   
   COP(M215_M1_DR_OUT_MAJ,M215_M1_DR_IN_MAJ,1);
   M215_M1_DR_IN_MAR.EN := M215_M1_DR_OUT_MAR.EN;
   M215_M1_DR_IN_MAR.PC := M215_M1_DR_OUT_MAR.PC;
   COP(M215_M1_DR_OUT_MAM,M215_M1_DR_IN_MAM,1);
   COP(M215_M1_DR_OUT_MAS,M215_M1_DR_IN_MAS,1);
   COP(M215_M1_DR_OUT_MRP,M215_M1_DR_IN_MRP,1);
   COP(M215_M1_DR_OUT_MCD,M215_M1_DR_IN_MCD,1);
   
   COP(M216_M1_DR_OUT_MAJ,M216_M1_DR_IN_MAJ,1);
   M216_M1_DR_IN_MAR.EN := M216_M1_DR_OUT_MAR.EN;
   M216_M1_DR_IN_MAR.PC := M216_M1_DR_OUT_MAR.PC;
   COP(M216_M1_DR_OUT_MAM,M216_M1_DR_IN_MAM,1);
   COP(M216_M1_DR_OUT_MAS,M216_M1_DR_IN_MAS,1);
   COP(M216_M1_DR_OUT_MRP,M216_M1_DR_IN_MRP,1);
   COP(M216_M1_DR_OUT_MCD,M216_M1_DR_IN_MCD,1);
   
   COP(M217_M1_DR_OUT_MAJ,M217_M1_DR_IN_MAJ,1);
   M217_M1_DR_IN_MAR.EN := M217_M1_DR_OUT_MAR.EN;
   M217_M1_DR_IN_MAR.PC := M217_M1_DR_OUT_MAR.PC;
   COP(M217_M1_DR_OUT_MAM,M217_M1_DR_IN_MAM,1);
   COP(M217_M1_DR_OUT_MAS,M217_M1_DR_IN_MAS,1);
   COP(M217_M1_DR_OUT_MRP,M217_M1_DR_IN_MRP,1);
   COP(M217_M1_DR_OUT_MCD,M217_M1_DR_IN_MCD,1);
   
   COP(M218_M1_DR_OUT_MAJ,M218_M1_DR_IN_MAJ,1);
   M218_M1_DR_IN_MAR.EN := M218_M1_DR_OUT_MAR.EN;
   M218_M1_DR_IN_MAR.PC := M218_M1_DR_OUT_MAR.PC;
   COP(M218_M1_DR_OUT_MAM,M218_M1_DR_IN_MAM,1);
   COP(M218_M1_DR_OUT_MAS,M218_M1_DR_IN_MAS,1);
   COP(M218_M1_DR_OUT_MRP,M218_M1_DR_IN_MRP,1);
   COP(M218_M1_DR_OUT_MCD,M218_M1_DR_IN_MCD,1);
   
   COP(M219_M1_DR_OUT_MAJ,M219_M1_DR_IN_MAJ,1);
   M219_M1_DR_IN_MAR.EN := M219_M1_DR_OUT_MAR.EN;
   M219_M1_DR_IN_MAR.PC := M219_M1_DR_OUT_MAR.PC;
   COP(M219_M1_DR_OUT_MAM,M219_M1_DR_IN_MAM,1);
   COP(M219_M1_DR_OUT_MAS,M219_M1_DR_IN_MAS,1);
   COP(M219_M1_DR_OUT_MRP,M219_M1_DR_IN_MRP,1);
   COP(M219_M1_DR_OUT_MCD,M219_M1_DR_IN_MCD,1);
   
   COP(M220_M1_DR_OUT_MAJ,M220_M1_DR_IN_MAJ,1);
   M220_M1_DR_IN_MAR.EN := M220_M1_DR_OUT_MAR.EN;
   M220_M1_DR_IN_MAR.PC := M220_M1_DR_OUT_MAR.PC;
   COP(M220_M1_DR_OUT_MAM,M220_M1_DR_IN_MAM,1);
   COP(M220_M1_DR_OUT_MAS,M220_M1_DR_IN_MAS,1);
   COP(M220_M1_DR_OUT_MRP,M220_M1_DR_IN_MRP,1);
   COP(M220_M1_DR_OUT_MCD,M220_M1_DR_IN_MCD,1);
   
   COP(M225_M1_DR_OUT_MAJ,M225_M1_DR_IN_MAJ,1);
   M225_M1_DR_IN_MAR.EN := M225_M1_DR_OUT_MAR.EN;
   M225_M1_DR_IN_MAR.PC := M225_M1_DR_OUT_MAR.PC;
   COP(M225_M1_DR_OUT_MAM,M225_M1_DR_IN_MAM,1);
   COP(M225_M1_DR_OUT_MAS,M225_M1_DR_IN_MAS,1);
   COP(M225_M1_DR_OUT_MRP,M225_M1_DR_IN_MRP,1);
   COP(M225_M1_DR_OUT_MCD,M225_M1_DR_IN_MCD,1);
   
END_ROUTINE

ROUTINE _101_LADDER   (* ladder *)
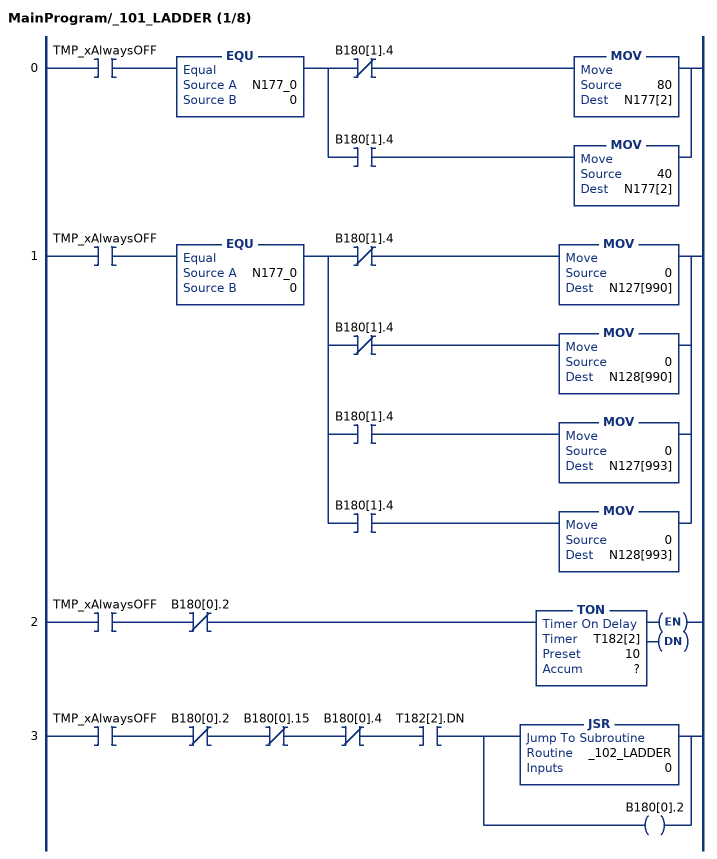
   0: XIC(TMP_xAlwaysOFF)EQU(N177_0,0)[XIO(B180[1].4) MOV(80,N177[2]) ,XIC(B180[1].4) MOV(40,N177[2]) ];
   1: XIC(TMP_xAlwaysOFF)EQU(N177_0,0)[XIO(B180[1].4) MOV(0,N127[990]) ,XIO(B180[1].4) MOV(0,N128[990]) ,XIC(B180[1].4) MOV(0,N127[993]) ,XIC(B180[1].4) MOV(0,N128[993]) ];
   2: XIC(TMP_xAlwaysOFF)XIO(B180[0].2)TON(T182[2],?,?);
   3: XIC(TMP_xAlwaysOFF)XIO(B180[0].2)XIO(B180[0].15)XIO(B180[0].4)XIC(T182[2].DN)[JSR(_102_LADDER,0) ,OTE(B180[0].2) ];
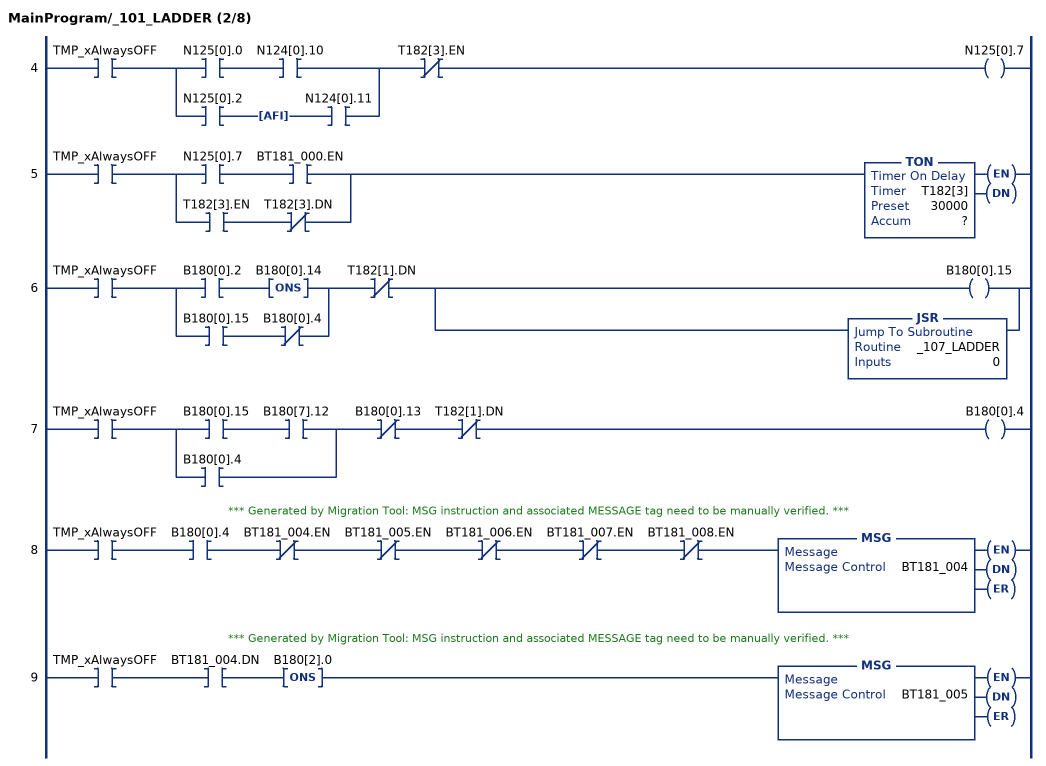
   4: XIC(TMP_xAlwaysOFF)[XIC(N125[0].0) XIC(N124[0].10) ,XIC(N125[0].2) AFI() XIC(N124[0].11) ]XIO(T182[3].EN)OTE(N125[0].7);
   5: XIC(TMP_xAlwaysOFF)[XIC(N125[0].7) XIC(BT181_000.EN) ,XIC(T182[3].EN) XIO(T182[3].DN) ]TON(T182[3],?,?);
   6: XIC(TMP_xAlwaysOFF)[XIC(B180[0].2) ONS(B180[0].14) ,XIC(B180[0].15) XIO(B180[0].4) ]XIO(T182[1].DN)[OTE(B180[0].15) ,JSR(_107_LADDER,0) ];
   7: XIC(TMP_xAlwaysOFF)[XIC(B180[0].15) XIC(B180[7].12) ,XIC(B180[0].4) ]XIO(B180[0].13)XIO(T182[1].DN)OTE(B180[0].4);
   // *** Generated by Migration Tool: MSG instruction and associated MESSAGE tag need to be manually verified. ***
   8: XIC(TMP_xAlwaysOFF)XIC(B180[0].4)XIO(BT181_004.EN)XIO(BT181_005.EN)XIO(BT181_006.EN)XIO(BT181_007.EN)XIO(BT181_008.EN)MSG(BT181_004);
   // *** Generated by Migration Tool: MSG instruction and associated MESSAGE tag need to be manually verified. ***
   9: XIC(TMP_xAlwaysOFF)XIC(BT181_004.DN)ONS(B180[2].0)MSG(BT181_005);
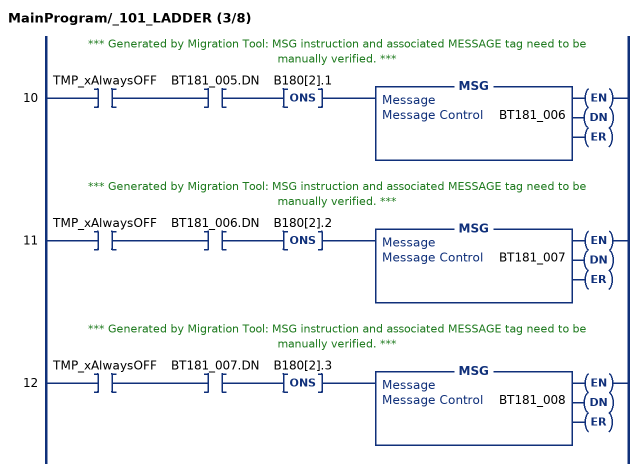
   // *** Generated by Migration Tool: MSG instruction and associated MESSAGE tag need to be manually verified. ***
   10: XIC(TMP_xAlwaysOFF)XIC(BT181_005.DN)ONS(B180[2].1)MSG(BT181_006);
   // *** Generated by Migration Tool: MSG instruction and associated MESSAGE tag need to be manually verified. ***
   11: XIC(TMP_xAlwaysOFF)XIC(BT181_006.DN)ONS(B180[2].2)MSG(BT181_007);
   // *** Generated by Migration Tool: MSG instruction and associated MESSAGE tag need to be manually verified. ***
   12: XIC(TMP_xAlwaysOFF)XIC(BT181_007.DN)ONS(B180[2].3)MSG(BT181_008);
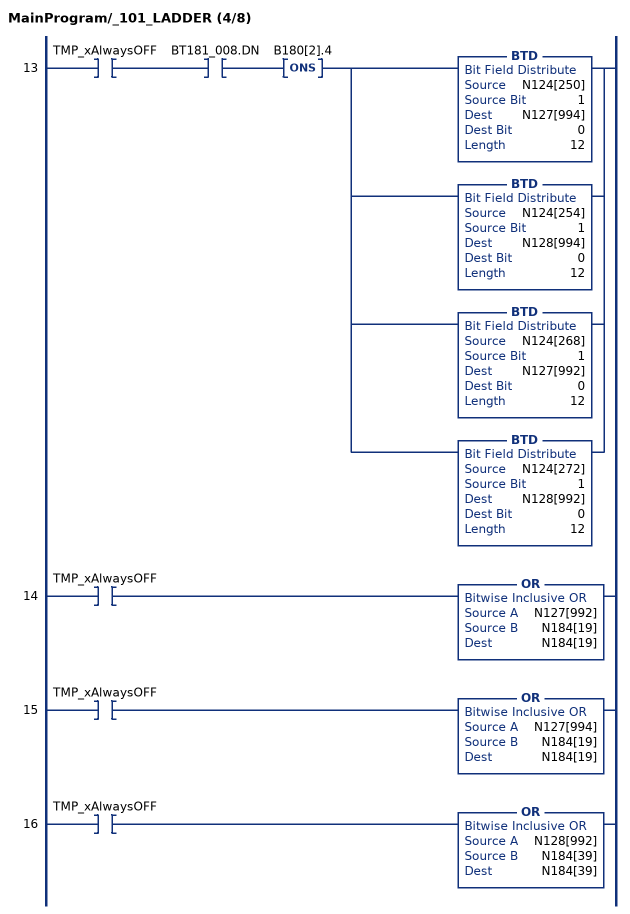
   13: XIC(TMP_xAlwaysOFF)XIC(BT181_008.DN)ONS(B180[2].4)[BTD(N124[250],1,N127[994],0,12) ,BTD(N124[254],1,N128[994],0,12) ,BTD(N124[268],1,N127[992],0,12) ,BTD(N124[272],1,N128[992],0,12) ];
   14: XIC(TMP_xAlwaysOFF)OR(N127[992],N184[19],N184[19]);
   15: XIC(TMP_xAlwaysOFF)OR(N127[994],N184[19],N184[19]);
   16: XIC(TMP_xAlwaysOFF)OR(N128[992],N184[39],N184[39]);
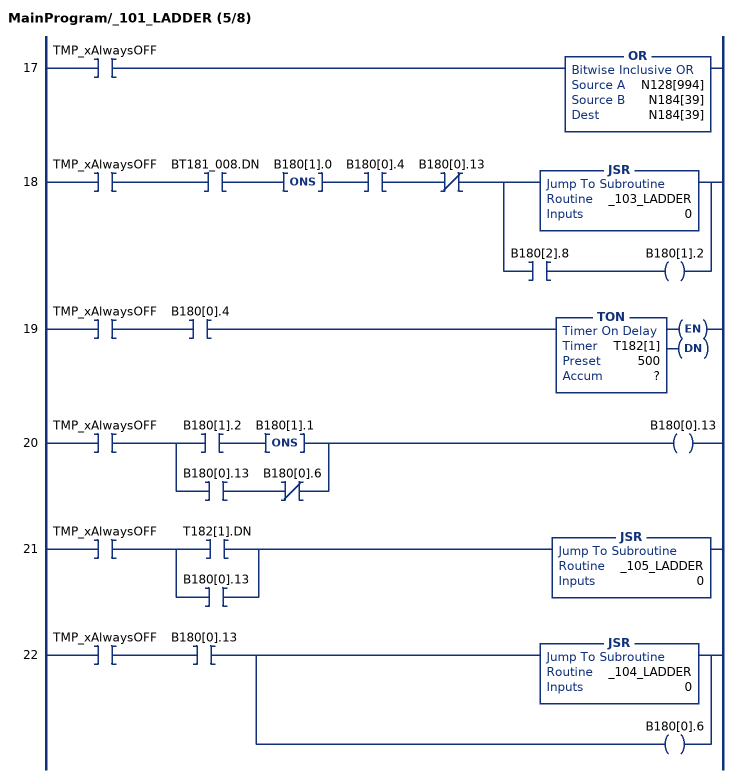
   17: XIC(TMP_xAlwaysOFF)OR(N128[994],N184[39],N184[39]);
   18: XIC(TMP_xAlwaysOFF)XIC(BT181_008.DN)ONS(B180[1].0)XIC(B180[0].4)XIO(B180[0].13)[JSR(_103_LADDER,0) ,XIC(B180[2].8) OTE(B180[1].2) ];
   19: XIC(TMP_xAlwaysOFF)XIC(B180[0].4)TON(T182[1],?,?);
   20: XIC(TMP_xAlwaysOFF)[XIC(B180[1].2) ONS(B180[1].1) ,XIC(B180[0].13) XIO(B180[0].6) ]OTE(B180[0].13);
   21: XIC(TMP_xAlwaysOFF)[XIC(T182[1].DN) ,XIC(B180[0].13) ]JSR(_105_LADDER,0);
   22: XIC(TMP_xAlwaysOFF)XIC(B180[0].13)[JSR(_104_LADDER,0) ,OTE(B180[0].6) ];
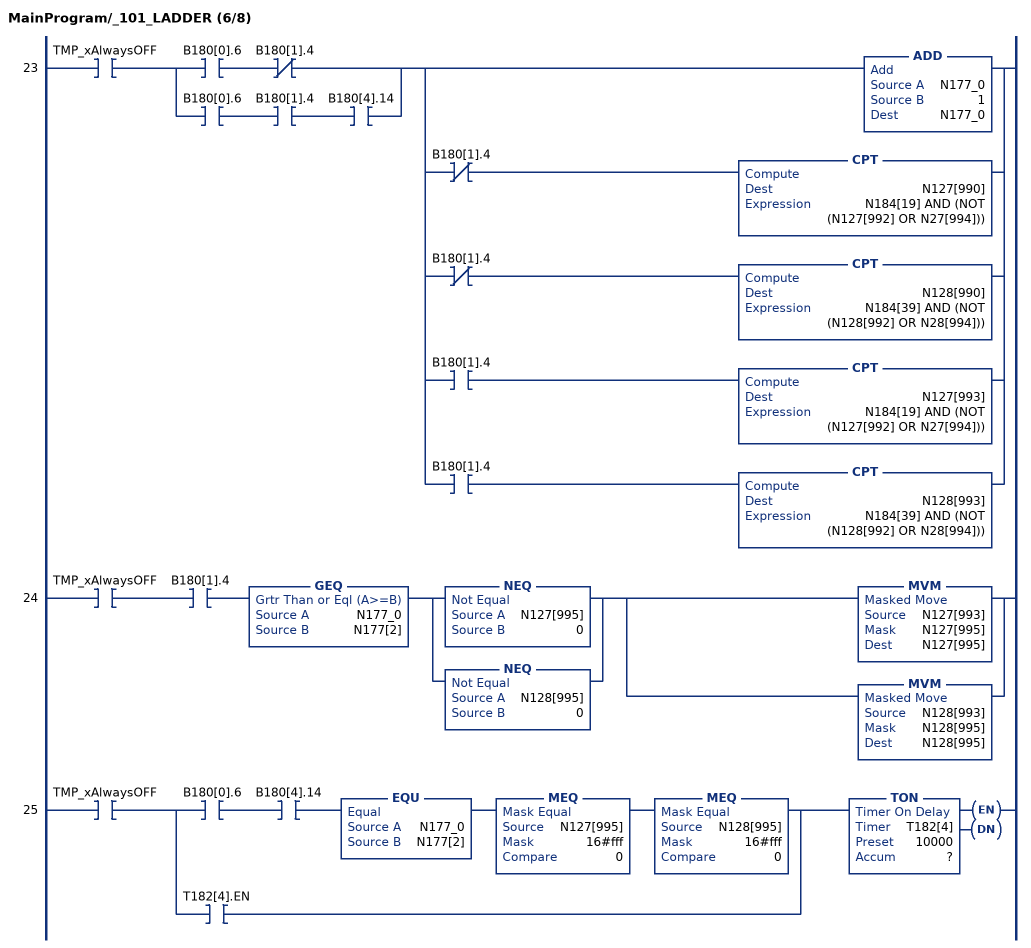
   23: XIC(TMP_xAlwaysOFF)[XIC(B180[0].6) XIO(B180[1].4) ,XIC(B180[0].6) XIC(B180[1].4) XIC(B180[4].14) ][ADD(N177_0,1,N177_0) ,XIO(B180[1].4) CPT(N127[990],N184[19] AND (NOT (N127[992] OR N27[994]))) ,XIO(B180[1].4) CPT(N128[990],N184[39] AND (NOT (N128[992] OR N28[994]))) ,XIC(B180[1].4) CPT(N127[993],N184[19] AND (NOT (N127[992] OR N27[994]))) ,XIC(B180[1].4) CPT(N128[993],N184[39] AND (NOT (N128[992] OR N28[994]))) ];
   24: XIC(TMP_xAlwaysOFF)XIC(B180[1].4)GEQ(N177_0,N177[2])[NEQ(N127[995],0) ,NEQ(N128[995],0) ][MVM(N127[993],N127[995],N127[995]) ,MVM(N128[993],N128[995],N128[995]) ];
   25: XIC(TMP_xAlwaysOFF)[XIC(B180[0].6) XIC(B180[4].14) EQU(N177_0,N177[2]) MEQ(N127[995],16#fff,0) MEQ(N128[995],16#fff,0) ,XIC(T182[4].EN) ]TON(T182[4],?,?);
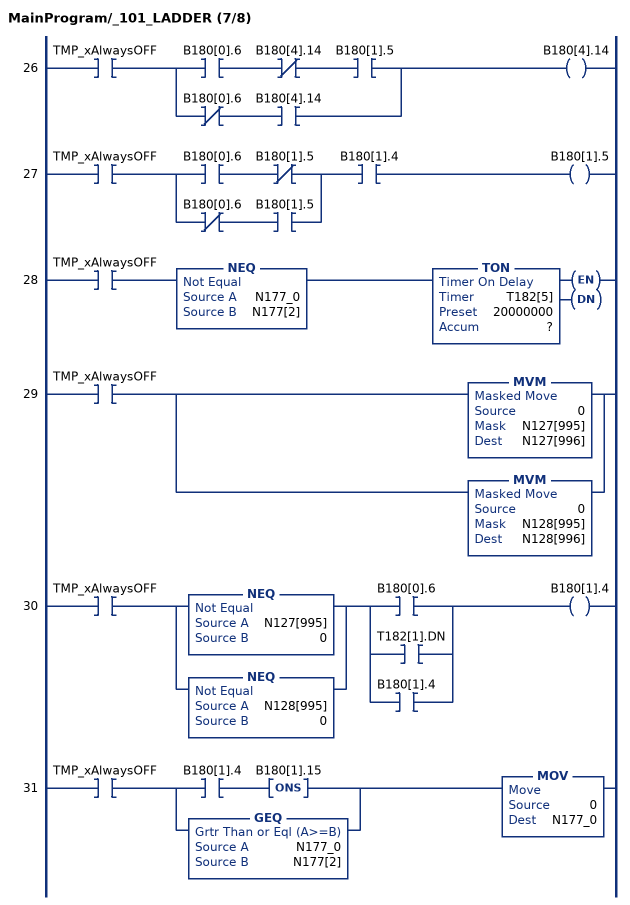
   26: XIC(TMP_xAlwaysOFF)[XIC(B180[0].6) XIO(B180[4].14) XIC(B180[1].5) ,XIO(B180[0].6) XIC(B180[4].14) ]OTE(B180[4].14);
   27: XIC(TMP_xAlwaysOFF)[XIC(B180[0].6) XIO(B180[1].5) ,XIO(B180[0].6) XIC(B180[1].5) ]XIC(B180[1].4)OTE(B180[1].5);
   28: XIC(TMP_xAlwaysOFF)NEQ(N177_0,N177[2])TON(T182[5],?,?);
   29: XIC(TMP_xAlwaysOFF)[MVM(0,N127[995],N127[996]) ,MVM(0,N128[995],N128[996]) ];
   30: XIC(TMP_xAlwaysOFF)[NEQ(N127[995],0) ,NEQ(N128[995],0) ][XIC(B180[0].6) ,XIC(T182[1].DN) ,XIC(B180[1].4) ]OTE(B180[1].4);
   31: XIC(TMP_xAlwaysOFF)[XIC(B180[1].4) ONS(B180[1].15) ,GEQ(N177_0,N177[2]) ]MOV(0,N177_0);
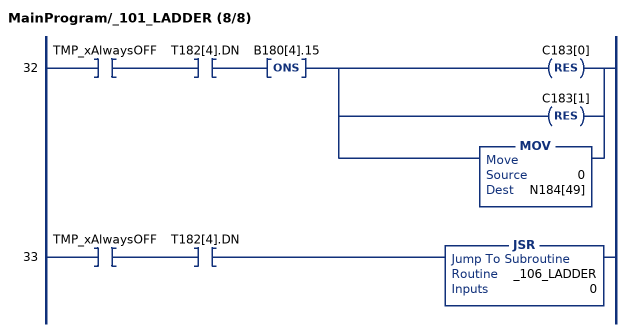
   32: XIC(TMP_xAlwaysOFF)XIC(T182[4].DN)ONS(B180[4].15)[RES(C183[0]) ,RES(C183[1]) ,MOV(0,N184[49]) ];
   33: XIC(TMP_xAlwaysOFF)XIC(T182[4].DN)JSR(_106_LADDER,0);
END_ROUTINE

ROUTINE _102_LADDER   (* ladder *)
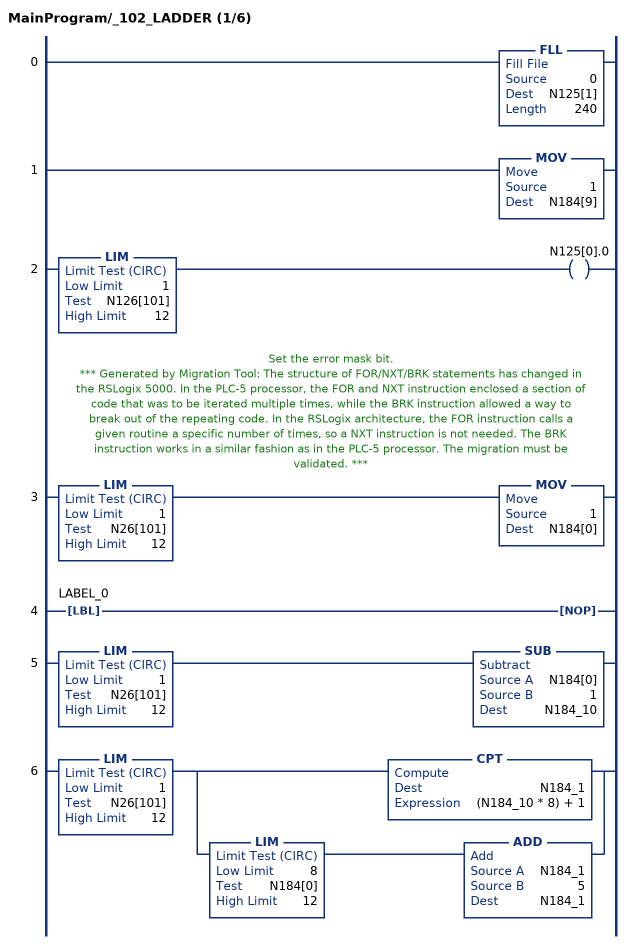
   0: FLL(0,N125[1],240);
   1: MOV(1,N184[9]);
   2: LIM(1,N126[101],12)OTE(N125[0].0);
   // Set the error mask bit.
   // *** Generated by Migration Tool: The structure of FOR/NXT/BRK statements has changed in the RSLogix 5000. In the PLC-5 processor, the FOR and NXT instruction enclosed a section of code that was to be iterated multiple times, while the BRK instruction allowed a way to break out of the repeating code. In the RSLogix architecture, the FOR instruction calls a given routine a specific number of times, so a NXT instruction is not needed. The BRK instruction works in a similar fashion as in the PLC-5 processor. The migration must be validated. ***
   3: LIM(1,N26[101],12)MOV(1,N184[0]);
   4: LBL(LABEL_0)NOP();
   5: LIM(1,N26[101],12)SUB(N184[0],1,N184_10);
   6: LIM(1,N26[101],12)[CPT(N184_1,(N184_10 * 8) + 1) ,LIM(8,N184[0],12) ADD(N184_1,5,N184_1) ];
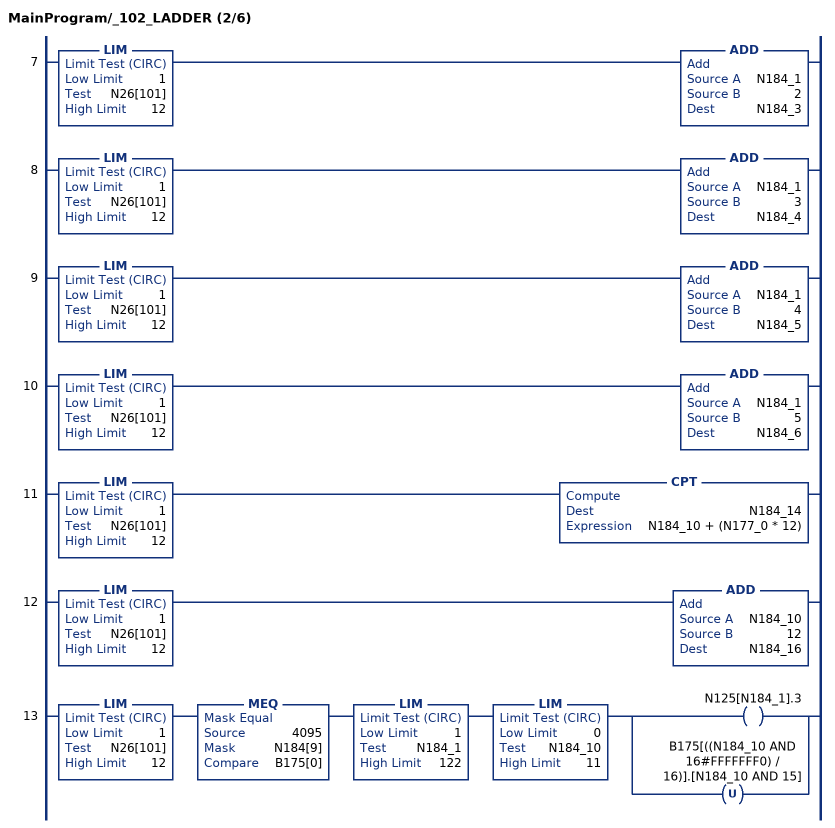
   7: LIM(1,N26[101],12)ADD(N184_1,2,N184_3);
   8: LIM(1,N26[101],12)ADD(N184_1,3,N184_4);
   9: LIM(1,N26[101],12)ADD(N184_1,4,N184_5);
   10: LIM(1,N26[101],12)ADD(N184_1,5,N184_6);
   11: LIM(1,N26[101],12)CPT(N184_14,N184_10 + (N177_0 * 12));
   12: LIM(1,N26[101],12)ADD(N184_10,12,N184_16);
   13: LIM(1,N26[101],12)MEQ(4095,N184[9],B175[0])LIM(1,N184_1,122)LIM(0,N184_10,11)[OTE(N125[N184_1].3) ,OTU(B175[((N184_10 AND 16#FFFFFFF0) / 16)].[N184_10 AND 15]) ];
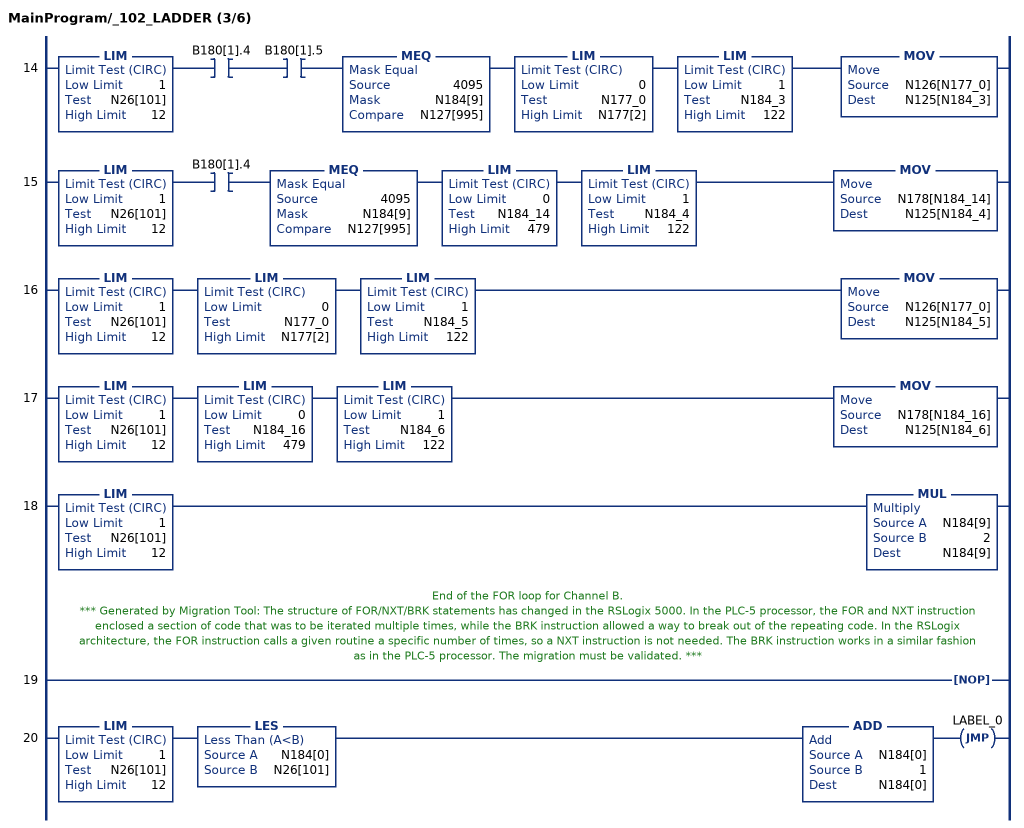
   14: LIM(1,N26[101],12)XIC(B180[1].4)XIC(B180[1].5)MEQ(4095,N184[9],N127[995])LIM(0,N177_0,N177[2])LIM(1,N184_3,122)MOV(N126[N177_0],N125[N184_3]);
   15: LIM(1,N26[101],12)XIC(B180[1].4)MEQ(4095,N184[9],N127[995])LIM(0,N184_14,479)LIM(1,N184_4,122)MOV(N178[N184_14],N125[N184_4]);
   16: LIM(1,N26[101],12)LIM(0,N177_0,N177[2])LIM(1,N184_5,122)MOV(N126[N177_0],N125[N184_5]);
   17: LIM(1,N26[101],12)LIM(0,N184_16,479)LIM(1,N184_6,122)MOV(N178[N184_16],N125[N184_6]);
   18: LIM(1,N26[101],12)MUL(N184[9],2,N184[9]);
   // End of the FOR loop for Channel B.
   // *** Generated by Migration Tool: The structure of FOR/NXT/BRK statements has changed in the RSLogix 5000. In the PLC-5 processor, the FOR and NXT instruction enclosed a section of code that was to be iterated multiple times, while the BRK instruction allowed a way to break out of the repeating code. In the RSLogix architecture, the FOR instruction calls a given routine a specific number of times, so a NXT instruction is not needed. The BRK instruction works in a similar fashion as in the PLC-5 processor. The migration must be validated. ***
   19: NOP();
   20: LIM(1,N26[101],12)LES(N184[0],N26[101])ADD(N184[0],1,N184[0])JMP(LABEL_0);
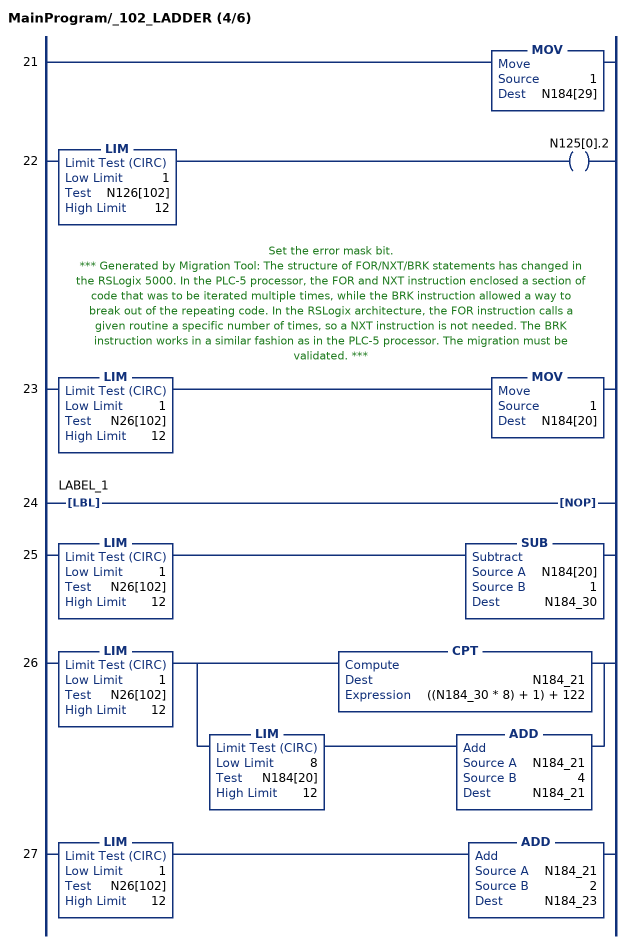
   21: MOV(1,N184[29]);
   22: LIM(1,N126[102],12)OTE(N125[0].2);
   // Set the error mask bit.
   // *** Generated by Migration Tool: The structure of FOR/NXT/BRK statements has changed in the RSLogix 5000. In the PLC-5 processor, the FOR and NXT instruction enclosed a section of code that was to be iterated multiple times, while the BRK instruction allowed a way to break out of the repeating code. In the RSLogix architecture, the FOR instruction calls a given routine a specific number of times, so a NXT instruction is not needed. The BRK instruction works in a similar fashion as in the PLC-5 processor. The migration must be validated. ***
   23: LIM(1,N26[102],12)MOV(1,N184[20]);
   24: LBL(LABEL_1)NOP();
   25: LIM(1,N26[102],12)SUB(N184[20],1,N184_30);
   26: LIM(1,N26[102],12)[CPT(N184_21,((N184_30 * 8) + 1) + 122) ,LIM(8,N184[20],12) ADD(N184_21,4,N184_21) ];
   27: LIM(1,N26[102],12)ADD(N184_21,2,N184_23);
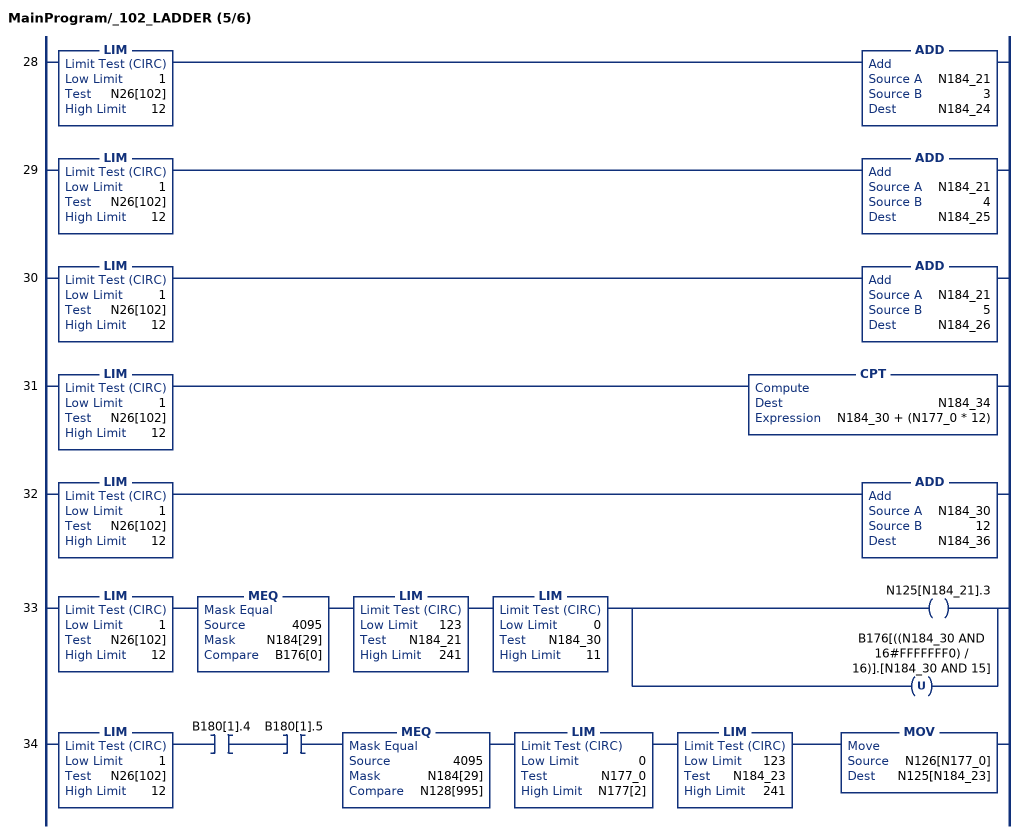
   28: LIM(1,N26[102],12)ADD(N184_21,3,N184_24);
   29: LIM(1,N26[102],12)ADD(N184_21,4,N184_25);
   30: LIM(1,N26[102],12)ADD(N184_21,5,N184_26);
   31: LIM(1,N26[102],12)CPT(N184_34,N184_30 + (N177_0 * 12));
   32: LIM(1,N26[102],12)ADD(N184_30,12,N184_36);
   33: LIM(1,N26[102],12)MEQ(4095,N184[29],B176[0])LIM(123,N184_21,241)LIM(0,N184_30,11)[OTE(N125[N184_21].3) ,OTU(B176[((N184_30 AND 16#FFFFFFF0) / 16)].[N184_30 AND 15]) ];
   34: LIM(1,N26[102],12)XIC(B180[1].4)XIC(B180[1].5)MEQ(4095,N184[29],N128[995])LIM(0,N177_0,N177[2])LIM(123,N184_23,241)MOV(N126[N177_0],N125[N184_23]);
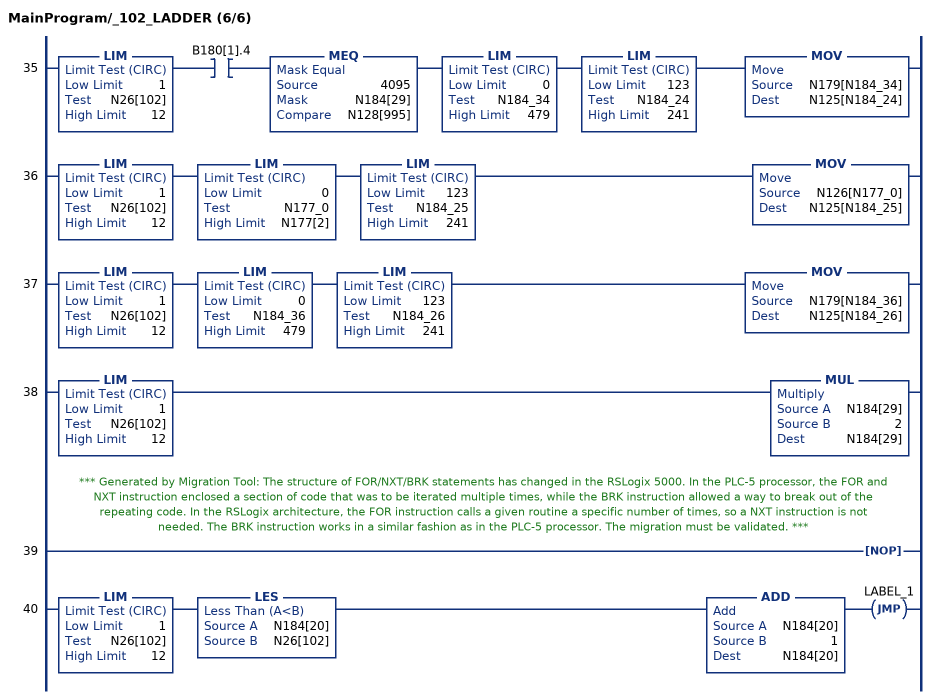
   35: LIM(1,N26[102],12)XIC(B180[1].4)MEQ(4095,N184[29],N128[995])LIM(0,N184_34,479)LIM(123,N184_24,241)MOV(N179[N184_34],N125[N184_24]);
   36: LIM(1,N26[102],12)LIM(0,N177_0,N177[2])LIM(123,N184_25,241)MOV(N126[N177_0],N125[N184_25]);
   37: LIM(1,N26[102],12)LIM(0,N184_36,479)LIM(123,N184_26,241)MOV(N179[N184_36],N125[N184_26]);
   38: LIM(1,N26[102],12)MUL(N184[29],2,N184[29]);
   // *** Generated by Migration Tool: The structure of FOR/NXT/BRK statements has changed in the RSLogix 5000. In the PLC-5 processor, the FOR and NXT instruction enclosed a section of code that was to be iterated multiple times, while the BRK instruction allowed a way to break out of the repeating code. In the RSLogix architecture, the FOR instruction calls a given routine a specific number of times, so a NXT instruction is not needed. The BRK instruction works in a similar fashion as in the PLC-5 processor. The migration must be validated. ***
   39: NOP();
   40: LIM(1,N26[102],12)LES(N184[20],N26[102])ADD(N184[20],1,N184[20])JMP(LABEL_1);
END_ROUTINE
